// Mitsubishi GX Works2 project: 20国轩1次注液出1031   PLC: Q06UDEH

TYPE ConveyorIO : STRUCT
  xUnloadCCW : BOOL;  (* 下料为反转 *)
  xUnloadAlarm : BOOL;  (* 下料报警 *)
  xUnload : BOOL;  (* 下料请求 *)
  xPutInto : BOOL;  (* 线体直接投入物料 *)
  xNotArriveAlarm : BOOL;  (* 未到达报警 *)
  xNextRun : BOOL;  (* 下段线体运行 *)
  xMotorCW : BOOL;  (* 电机正转 *)
  xMotorCCW : BOOL;  (* 电机反转 *)
  xManual : BOOL;  (* 手动 *)
  xloadCCW : BOOL;  (* 上料为反转 *)
  xLimitAlarrm : BOOL;  (* 限位报警 *)
  xLoad : BOOL;  (* 上料请求 *)
  xForward : BOOL;  (* 正转手动 *)
  xEmpty : BOOL;  (* 线体状态为空 *)
  xCWPresent : BOOL;  (* 正转检测有无传感器 *)
  xCCWPresent : BOOL;  (* 反转检测有无传感器 *)
  xBusy : BOOL;  (* 工作中 *)
  xBackward : BOOL;  (* 反转手动 *)
  xAuto : BOOL;  (* 自动 *)
  xPosLimit : BOOL;  (* 正限位 *)
  xNegLimit : BOOL;  (* 负限位 *)
  xOverWidthAlarm : BOOL;  (* 超宽报警 *)
  xError : BOOL;  (* 报警 *)
  iProductCategoryIn : INT;  (* 产品类型输入 *)
  iProductCategory : INT;  (* 产品类型记录 *)
  iProductCategoryOut : INT;  (* 产品类型输出 *)
  diDeviceID : DINT;  (* 设备编号 *)
  tUnloadAlarmDelay : TIME;  (* 下料报警时间设置 *)
  tLoadDelay : TIME;  (* 上料延时设置 *)
  xSizeDeficientDetect : BOOL;  (* 尺寸缺陷检测 *)
  xZoneClear : BOOL;  (* 初始化线体清除 *)
  tZoneClearTime : TIME;  (* 初始化线体清除时间 *)
  iTaskIDIn : INT;  (* 产品类型输入 *)
  iTaskID : INT;  (* 产品类型记录 *)
  iTaskIDOut : INT;  (* 产品类型输出 *)
  diDesConveyorIn : DINT;  (* 产品类型输入 *)
  diDesConveyor : DINT;  (* 产品类型记录 *)
  diDesConveyorOut : DINT;  (* 产品类型输出 *)
END_STRUCT END_TYPE

TYPE QueueElement : STRUCT
  xCondition : BOOL;
  iPriority : INT;
END_STRUCT END_TYPE

TYPE ShuttleCarIO : STRUCT
  xReady : BOOL;  (* 准备就绪 *)
  xForward : BOOL;  (* 正转 *)
  xBackward : BOOL;  (* 反转 *)
  iCurrentPos : INT;  (* 当前位置 *)
  iDestinationPos : INT;  (* 目标位置 *)
  xCW : BOOL;  (* 正转输出 *)
  xCCW : BOOL;  (* 反转输出 *)
  xBrake : BOOL;  (* 刹车 *)
  xHomeSwitch : BOOL;  (* 零位接近开关 *)
  xPosLimit : BOOL;  (* 正限位 *)
  xNegLimit : BOOL;  (* 负限位 *)
  xMDIExe : BOOL;  (* MDI开始 *)
  xMDIDone : BOOL;  (* MDI 完成 *)
  xPassLimit : BOOL;  (* 限位屏蔽 *)
  xPosLimitCatch : BOOL;  (* 正限位捕捉 *)
  xNegLimitCatch : BOOL;  (* 负限位捕捉 *)
  xHomeExe : BOOL;  (* 开始寻零 *)
  xHomeDone : BOOL;  (* 寻零完成 *)
  xHomeBusy : BOOL;  (* 寻零中 *)
  xHomeFailed : BOOL;  (* 寻零失败 *)
  xBusy : BOOL;  (* 工作中 *)
  tArriveDelay : TIME;  (* 到位延时 *)
  xCylinder : BOOL;  (* 气缸控制 *)
  tBrakeDelay : TIME;  (* 抱闸延时 *)
  xPauseRamp : BOOL;  (* 暂停减速斜坡标志位 *)
  xPresentDetect1 : BOOL;  (* 物料有无检测1 *)
  xPresentDetect2 : BOOL;  (* 物料有无检测2 *)
  xOvertimeAlarm : BOOL;  (* 超时报警 *)
  tSetOverTime : TIME;  (* 设置超时时间 *)
  xLooseDetect : BOOL;  (* 松绳检测 *)
  xLooseAlarm : BOOL;  (* 松绳报警 *)
  xArrive : BOOL;  (* 到位信号 *)
  diDeviceID : DINT;  (* 设备编号 *)
  xMoveStep : BOOL;  (* 寸动 *)
  xAdrSwitch : ARRAY [1..8] OF BOOL;  (* 位置开关 *)
END_STRUCT END_TYPE

TYPE SwitchIO : STRUCT
  xLiftCylinderRetractDetect : BOOL;
  xLiftCylinderExtendDetect : BOOL;
  xLiftCylinderRetract : BOOL;
  xLiftCylinderExtend : BOOL;
  xEntryBarCylinderRetract : BOOL;
  xLiftCylinderExtendInit : BOOL;
  xEntryEnable : BOOL;
  xExitEnable : BOOL;
  xExitBarCylinderRetract : BOOL;
  xSwithEnable : BOOL;
  xLiftCylinderRetractButton : BOOL;
  xLiftCylinderExtendButton : BOOL;
  xEntryBarCylinderRetractButton : BOOL;
  xExitBarCylinderRetractButton : BOOL;
  xPutInto : BOOL;  (* 单体复位 *)
  tSetOvertime : TIME;  (* 设定超时报警时间 *)
  xOvertimeAlarm : BOOL;  (* 超时报警 *)
END_STRUCT END_TYPE

TYPE UConveyorIO : STRUCT
  xLiftCylinderRetractDetect1 : BOOL;
  xLiftCylinderRetractDetect2 : BOOL;
  xLiftCylinderExtendDetect1 : BOOL;
  xLiftCylinderExtendDetect2 : BOOL;
  xLiftCylinderRetract1 : BOOL;
  xLiftCylinderRetract2 : BOOL;
  xLiftCylinderExtend1 : BOOL;
  xLiftCylinderExtend2 : BOOL;
  xExitBarCylinderRetract1 : BOOL;
  xExitBarCylinderRetract2 : BOOL;
  xLiftCylinderExtendInit1 : BOOL;
  xLiftCylinderExtendInit2 : BOOL;
  xEntryEnable1 : BOOL;
  xEntryEnable2 : BOOL;
  xEntryEnable3 : BOOL;
  xExitEnable1 : BOOL;
  xExitEnable2 : BOOL;
  xExitEnable3 : BOOL;
  xPassEnable : BOOL;  (* 直接放行去下段 *)
  xLiftCylinderRetractButton1 : BOOL;
  xLiftCylinderRetractButton2 : BOOL;
  xLiftCylinderExtendButton1 : BOOL;
  xLiftCylinderExtendButton2 : BOOL;
  xExitBarCylinderRetractButton1 : BOOL;
  xExitBarCylinderRetractButton2 : BOOL;
  xPutInto : BOOL;  (* 单体复位 *)
  tSetOvertime : TIME;  (* 设定超时报警时间 *)
  xOvertimeAlarm : BOOL;  (* 超时报警 *)
  iTask : INT;  (* 3个任务 *)
  xBatteryDetect1 : BOOL;  (* 电池检测1 *)
  xBatteryDetect2 : BOOL;  (* 电池检测2 *)
  xBatteryError : BOOL;  (* 空框里有电池错误 *)
END_STRUCT END_TYPE

TYPE FanucRobotIO : STRUCT
  i_xCMDENBL : BOOL;
  i_xSYSRDY : BOOL;
  i_xPROG_RUN : BOOL;  (* 程序运行中 *)
  i_xPAUSED : BOOL;
  i_xHELD : BOOL;
  i_xFAULT : BOOL;
  i_xATPERCH : BOOL;
  i_xTPENBL : BOOL;
  i_xBATALM : BOOL;
  i_xBUSY : BOOL;  (* 工作中信号 *)
  i_arrxSNO : ARRAY [0..7] OF BOOL;  (* 传回的数据 *)
  i_xSNACK : BOOL;  (* 数据传回校验标志位 *)
  o_xIMSTP : BOOL;
  o_xHOLD : BOOL;
  o_xSFSPD : BOOL;
  o_xCSTOPI : BOOL;
  o_xRESET : BOOL;
  o_xSTART : BOOL;
  o_xENBL : BOOL;
  o_iPNS : INT;  (* 发给他的动作编号 *)
  o_xPNSTROBE : BOOL;  (* 传递动作编号标志位 *)
  o_xPROD_START : BOOL;  (* 启动信号，下降沿开动 *)
  o_xREMOTE : BOOL;  (* 远程模式开启 *)
  i_xCommandStart : BOOL;  (* 启动 *)
  i_iMotionNumber : INT;  (* 我程序给的动作编号 *)
  o_xPNSFailed : BOOL;  (* 程序号传输错误 *)
  o_uiOffset_X : INT;  (* X轴偏移量 *)
  o_uiOffset_Y : INT;  (* Y轴偏移量 *)
  io_xMutexLock : BOOL;  (* 互斥锁 *)
END_STRUCT END_TYPE

TYPE CommunicationIO : STRUCT
  i_iResponsPCPLC : INT;  (* 上位机写入-请求确认 *)
  i_iReadWriteFlagPCPLC : INT;  (* 上位机写入-读写标志位 *)
  i_iTaskProcessFlagPCPLC : INT;  (* 上位机写入-任务出料标志位 *)
  i_iCommandPCPLC : INT;  (* 上位机写入-命令字 *)
  i_iTaskIDPCPLC : INT;  (* 上位机写入-任务号 *)
  i_diDestinationDevicePCPLC : DINT;  (* 上位机写入-目标设备号 *)
  i_iProductIDPCPLC : INT;  (* 上位机写入-框码后4位 *)
  o_iRequestPLCPC : INT;  (* 上位机读取-请求状态 *)
  o_iReadWriteFlagPLCPC : INT;  (* 上位机读取-读写标志位 *)
  o_iDeviceStatusPLCPC : INT;  (* 上位机读取-设备状态 *)
  o_iTaskIDPLCPC : INT;  (* 上位机读取-任务号 *)
  o_iProductIDPLCPC : INT;  (* 上位机读取-框码后4位 *)
END_STRUCT END_TYPE

TYPE PackCommunicationIO : STRUCT
  i_iResponsPCPLC : INT;  (* 上位机写入-请求确认 *)
  i_iPackDoneAknPCPLC : INT;  (* 上位机写入-放行 *)
  i_iSinglePackResponsePCPLC : INT;  (* 上位机写入-单次装载应答 *)
  i_iSinglePackDoneAknPCPLC : INT;  (* 上位机写入-单次装载处理完成 *)
  o_iRequestPLCPC : INT;  (* 上位机读取-装载请求 *)
  o_iPackDonePLCPC : INT;  (* 上位机读取-装载完成 *)
  o_iSinglePackRequestPLCPC : INT;  (* 上位机读取-单次装载请求 *)
  o_iSinglePackDonePLCPC : INT;  (* 上位机读取-单次装载完成 *)
  o_iXCoordinatePLCPC : INT;  (* 上位机读取-行坐标 *)
  o_iYCoordinatePLCPC : INT;  (* 上位机读取-列坐标 *)
  o_arrwCode : ARRAY [0..7] OF BOOL;  (* 上位机读取-电芯码 *)
END_STRUCT END_TYPE

TYPE BatteryCode : STRUCT
  arrwCode : ARRAY [0..8] OF WORD;
END_STRUCT END_TYPE

// global labels: Global
VAR_GLOBAL
  g_xAuto AT M11 : BOOL;
  g_xManual : BOOL;
  g_xEStop AT X0 : BOOL;
  g_xReset AT X4 : BOOL;
  g_xStackLampRed AT Y200 : BOOL;
  g_xStackLampAmber AT Y201 : BOOL;
  g_xStackLampGreen AT Y202 : BOOL;
  g_xBuzzer AT Y203 : BOOL;
  g_xStop AT X3 : BOOL;
  g_xAutoStart AT X2 : BOOL;
  g_xRemoteAutoStart AT M0 : BOOL;
  g_xRemoteAuto AT M10 : BOOL;
  g_iState AT D40 : INT;
  g_iLocalAutoStep : BOOL;
  g_xAlarm : BOOL;
  g_xPause AT M3 : BOOL;  (* 暂停 *)
  g_diDeviceIDSelect AT D0 : DINT;
  g_xResetSingle AT M4 : BOOL;  (* 单线体复位 *)
  g_xInsertTask AT M5 : BOOL;  (* 插入任务 *)
  g_iInsertTaskID AT D2 : INT;  (* 插入任务号 *)
  g_iConveyorStatus AT D4 : INT;
  g_iInsertCategory AT D6 : INT;
  g_diInsertDesConveyor AT D8 : DINT;
  g_xTcpFailed : BOOL;
  g_xPickOver : ARRAY [1..4] OF BOOL;  (* 注液机给我们的信号，待定 *)
  g_xRobot1BatteryDetect : ARRAY [1..8] OF BOOL;
  g_xRobot2BatteryDetect : ARRAY [1..8] OF BOOL;
  g_xRobot3BatteryDetect : ARRAY [1..8] OF BOOL;
  g_xRobot4BatteryDetect : ARRAY [1..8] OF BOOL;
  g_xAutoLamp AT Y204 : BOOL;
  g_xAutoSwitch AT X1 : BOOL;
  g_xMute : BOOL;
  g_iLoadTask AT D50 : ARRAY [0..13] OF INT;
  g_xResetTask1 AT M9 : BOOL;  (* 复位排队任务的 *)
END_VAR

// global labels: Pro
VAR_GLOBAL
  g_xRobot1Pos1Done AT X0A0 : BOOL;  (* 机器人1工位1码垛完成 *)
  g_xRobot1Pos1Ready AT Y230 : BOOL;  (* 机器人1工位1空托盘到位 *)
  g_xRobot1Pos2Done AT X0A1 : BOOL;  (* 机器人1工位2码垛完成 *)
  g_xRobot1Pos2Ready AT Y231 : BOOL;  (* 机器人1工位2空托盘到位 *)
  g_xRobot2Pos1Done AT X0A2 : BOOL;  (* 机器人2工位1码垛完成 *)
  g_xRobot2Pos1Ready AT Y237 : BOOL;  (* 机器人2工位1空托盘到位 *)
  g_xRobot2Pos2Done AT X0A3 : BOOL;  (* 机器人2工位2码垛完成 *)
  g_xRobot2Pos2Ready AT Y239 : BOOL;  (* 机器人2工位2空托盘到位 *)
  g_xRobot3Pos1Done AT X0A4 : BOOL;  (* 机器人3工位1码垛完成 *)
  g_xRobot3Pos1Ready AT Y232 : BOOL;  (* 机器人3工位1空托盘到位 *)
  g_xRobot3Pos2Done AT X0A5 : BOOL;  (* 机器人3工位2码垛完成 *)
  g_xRobot3Pos2Ready AT Y233 : BOOL;  (* 机器人3工位2空托盘到位 *)
  g_xRobot4Pos1Done AT X0A6 : BOOL;  (* 机器人4工位1码垛完成 *)
  g_xRobot4Pos1Ready : BOOL;  (* 机器人4工位1空托盘到位 *)
  g_xRobot4Pos2Done AT X0A7 : BOOL;  (* 机器人4工位2码垛完成 *)
  g_xRobot4Pos2Ready : BOOL;  (* 机器人4工位2空托盘到位 *)
END_VAR

// task Task_01 (event TRUE, interval 0, priority 31): POU, TCP, START

FUNCTION_BLOCK Conveyor
VAR
  m_xPresentDelay : BOOL;  (* 有无判断延时 *)
  m_xLoadDelayOut : BOOL;  (* 上料延时输出 *)
  m_xInitial : BOOL;  (* 初始化 *)
  m_tUnloadTimer : TIME;  (* 下料计时器 *)
  m_tPresentDelayCurrentTime : TIME;
  m_tonUnloadAlam : TON;  (* 下料报警定时器 *)
  m_tonPresentDelay : TON;  (* 物料有无判断延时，防止误动作 *)
  m_tonNotArriveAlarm : TON;  (* 未到达报警计时 *)
  m_tonLoadDelay : TON;  (* 上料延时 *)
  m_tNotArriveCurrentTime : TIME;  (* 未到达报警计时当前时间 *)
  m_tLoadTimer : TIME;  (* 上料计时器 *)
  iStep : INT;  (* 上料步骤 *)
  m_wStateWord : INT;
END_VAR
VAR_IN_OUT
  ConveyorMotor : ConveyorIO;  (* 输送线输入输出 *)
END_VAR
VAR
  m_tonZoneClear : TON;  (* 初始化清除 *)
  m_tZoneClearCurrentTime : TIME;  (* 初始化清除当前时间 *)
  m_xAutoClear : BOOL;  (* 初始化清除标志位 *)
  m_xZoneClearDone : BOOL;  (* 初始化清除完成 *)
END_VAR
(*////////////////////////////////////////////////////////////////////////////////////////////////////////////
//传输线控制FB块，可控制单方向线体，双向旋转线体，支持双向上下料            
//线体初始化后为空的情况下输入xLoad信号即可进行上料动作，使用xLoadCCW信号可反方向上料
//增加了产品信息和产品种类的储存，当传输线为空和上料进行标志位为零的情况下清除产品信息和产品种类
//使用方式是在置位xLoad信号后，把产品信息和产品种类传入，等下料后自动清零
//线体不为空的情况下使用xUnload信号可进行下料动作，物料有无传感器的下降沿后出发计时器，延时断开传输线旋转
//单方向传输线体把xLoadCCW、xUnloadCCW设置为零，双向线体上料方向和下料反向的,方向固定的 把xUnloadCCW设置为1
//双方向线体双向都能上下料的要根据上料的方向来设置xLoadCCW,xUnloadCCW
//增加工作中信号xBusy当电机正转 显示为工作中
//增加上下料超时报警，xLoadAlarm，xUnloadAlarm，设定时间在LOAD_UNLOAD_TIME常量上，现在设置的为30秒
//增加xPutInto信号，用于直接投入的物料，检测开关感应到后，直接进入下料流程，上升沿有效
//离开延时改为变量 iLeaveDelay 默认为0 离开检测开关离输送线尾端比较远的线体需要根据情况设定100ms为单位
//增加初始化标志位，增加进入延时时间，初始化为进入延时时间为0 ，离开延时时间为2S，通过外围接口可以更改
//修改信息  修改后请增加版本
//12-17进行了优化，增加了未到达报警，当物料未传送到下一设备，就报未到达报警，使用xNextRun标志位制作，没有正常到达
//第0步，不能跳转到第一步把标志位复位，即出现中断情况，2秒后报警
//修改信息  修改后请增加版本
//上料延时增加为50ms防止干扰信号
//nextrun信号在 第三步也要复位
//增加限位报警
//增加超宽报警
//增加产品型号输出在下料的时候把产品型号输送给下一段线体
//增加线体单独复位
//增加任务插入功能配合全局变量
//增加暂停功能
//增加线体状态字显示  0 空闲 1：有料  2 工作中  3  超限报警 4 超宽报警  5 未到达报警  6 下料超时报警
//空料判断放在自动前，进行有无报警判断，然后跳转
//修改超限报警，与尺寸检测报警
////YAO      V1.0
//把所有的IF语句去掉，  IF语句占用指针存储区，容易造成存储区不足的现象
////YAO      V1.1
//初始化清除线体标志位xZoneClear
//ZPA zero pressure accumulation  Term that describes the Conveyor controls and mechanical scheme that will 
//cause loads to queue on a conveyor in discrete zones such that loads do not touch each other(wrapped boxed tray tote carton)
//除了产品信息外，还增加了目标地址，任务类型的数据传递。
//YAO      V1.0
///////////////////////////////////////////////////////////////////////////////////////////////////////////
(*********************************************************)
(*//初始化，
//上料延时位0S，下料报警延时为30S
//下料延时设一个比较大的时间，主要依靠xunload标志位来停止输送线，特殊情况可以用延时来停止物流线下料
//设置时间大的时候计时器会失效*)
IF NOT m_xInitial THEN
	ConveyorMotor.tLoadDelay:=T#100ms;
	ConveyorMotor.tUnloadAlarmDelay:=T#30s;
	ConveyorMotor.xPosLimit:=1;
	ConveyorMotor.xNegLimit:=1;
	ConveyorMotor.xSizeDeficientDetect:=0;
	ConveyorMotor.xZoneClear:=0;
	ConveyorMotor.tZoneClearTime:=T#10s;
	m_xInitial:=1;
END_IF;
(*//自动
//复位信号把步号置0，但xLoad与xUnload没有复位，调用程序需要注意复位后把这两个信号置零，以免发生误动作
//物料有无判断增加延时，防止开自动瞬间误动作发生*)
m_tonPresentDelay(IN:= ConveyorMotor.xCWPresent OR ConveyorMotor.xCCWPresent,
 PT:=T#100ms,
 Q:= m_xPresentDelay,
 ET:= m_tPresentDelayCurrentTime);
CASE iStep OF
0:(*//初始化*)
	ConveyorMotor.xMotorCW:=0;
	ConveyorMotor.xMotorCCW:=0;
	ConveyorMotor.xNextRun:=0;
	ConveyorMotor.iProductCategoryOut:=0;
	ConveyorMotor.iTaskIDOut:=0;
	ConveyorMotor.diDesConveyorOut:=0;
	out(NOT m_xPresentDelay,ConveyorMotor.xEmpty);(*	//判断物料有无传感器*)	
	mov(m_xPresentDelay AND g_xAuto AND NOT ConveyorMotor.xError,3,iStep);(*//自动情况下进行跳转*)(*无超限报警*)
	mov(NOT m_xPresentDelay AND g_xAuto AND NOT ConveyorMotor.xError,1,iStep);
1: (*//上料*)
	rst(ConveyorMotor.xLoad ,ConveyorMotor.iProductCategory);(*//上料开始清除产品信息*)
	rst(ConveyorMotor.xLoad ,ConveyorMotor.iTaskID);
	rst(ConveyorMotor.xLoad ,ConveyorMotor.diDesConveyor);
	mov(ConveyorMotor.xLoad,2,iStep);
2: (*//上料完成*)
	ConveyorMotor.iProductCategory:=ConveyorMotor.iProductCategoryIn;(* //产品信息传入*)
	ConveyorMotor.iTaskID:=ConveyorMotor.iTaskIDIn;
	ConveyorMotor.diDesConveyor:=ConveyorMotor.diDesConveyorIn;
	set(ConveyorMotor.xloadCCW,ConveyorMotor.xMotorCCW);
	rst(ConveyorMotor.xloadCCW,ConveyorMotor.xMotorCW);
	set(NOT ConveyorMotor.xloadCCW,ConveyorMotor.xMotorCW);
	rst(NOT ConveyorMotor.xloadCCW,ConveyorMotor.xMotorCCW);	
	m_tonLoadDelay(IN:= (ConveyorMotor.xCWPresent AND NOT ConveyorMotor.xloadCCW) 
  		OR (ConveyorMotor.xCCWPresent AND ConveyorMotor.xloadCCW) ,
  PT:= ConveyorMotor.tLoadDelay ,
  Q:= m_xLoadDelayOut ,
  ET:= m_tLoadTimer );
	mov(m_xLoadDelayOut,3, iStep);
3:(*//下料请求*)	
	ConveyorMotor.xMotorCW:=0;
	ConveyorMotor.xMotorCCW:=0;
	ConveyorMotor.xEmpty:=0;
	mov(ConveyorMotor.xUnload AND NOT ConveyorMotor.xOverWidthAlarm,4,iStep);
4:(*	//下料完成*)
	set(ConveyorMotor.xUnloadCCW,ConveyorMotor.xMotorCCW);
	rst(ConveyorMotor.xUnloadCCW,ConveyorMotor.xMotorCW);
	set(NOT ConveyorMotor.xUnloadCCW,ConveyorMotor.xMotorCW);
	rst(NOT ConveyorMotor.xUnloadCCW,ConveyorMotor.xMotorCCW);	
	ConveyorMotor.xNextRun:=1; (*下一段线体旋转*)
	ConveyorMotor.iProductCategoryOut:=ConveyorMotor.iProductCategory;(*产品型号输出给下一段线体*)
	ConveyorMotor.iTaskIDOut:=ConveyorMotor.iTaskID;
	ConveyorMotor.diDesConveyorOut:=ConveyorMotor.diDesConveyor;
	mov( NOT ConveyorMotor.xUnload , 0, istep );
END_CASE;
(*In-feed zone clear and ready to accept a load from upstream Conveyor*)
set(ldp(TRUE,g_xAuto) ,m_xAutoClear);
rst(ldf(TRUE,g_xAuto) ,m_xAutoClear);
m_tonZoneClear(IN:= m_xAutoClear AND ConveyorMotor.xZoneClear ,PT:= ConveyorMotor.tZoneClearTime ,Q:=m_xZoneClearDone ,ET:= m_tZoneClearCurrentTime );
set(m_xAutoClear AND ConveyorMotor.xZoneClear,ConveyorMotor.xMotorCW);
mov( m_xAutoClear AND ConveyorMotor.xZoneClear, 0 ,iStep );
rst(  ldf(TRUE, m_xAutoClear ) ,ConveyorMotor.xMotorCW);
rst( m_xZoneClearDone OR m_xPresentDelay  , m_xAutoClear );
(*投入上料，搬出下料，也可用来初始化*)
movp( ConveyorMotor.xPutInto, 0 , iStep );
(*//当前任务显示*)
movp( ConveyorMotor.diDeviceID=g_diDeviceIDSelect , ConveyorMotor.iProductCategory , g_iInsertCategory );
movp( ConveyorMotor.diDeviceID=g_diDeviceIDSelect , ConveyorMotor.iTaskID , g_iInsertTaskID );
dmovp( ConveyorMotor.diDeviceID=g_diDeviceIDSelect , ConveyorMotor.diDesConveyor , g_diInsertDesConveyor );
(*//插入任务*)
mov(g_xInsertTask AND ConveyorMotor.diDeviceID=g_diDeviceIDSelect ,g_iInsertCategory , ConveyorMotor.iProductCategory );
mov(g_xInsertTask AND ConveyorMotor.diDeviceID=g_diDeviceIDSelect , g_iInsertTaskID , ConveyorMotor.iTaskID );
dmov(g_xInsertTask AND ConveyorMotor.diDeviceID=g_diDeviceIDSelect , g_diInsertDesConveyor , ConveyorMotor.diDesConveyor );
(*//单线体复位，当设备号与本线体一致的时候执行复位*)
mov(g_xResetSingle AND ConveyorMotor.diDeviceID=g_diDeviceIDSelect , 0 , iStep );
rst(g_xResetSingle AND ConveyorMotor.diDeviceID=g_diDeviceIDSelect ,ConveyorMotor.xNextRun );
rst(g_xResetSingle AND ConveyorMotor.diDeviceID=g_diDeviceIDSelect  ,ConveyorMotor.xLimitAlarrm );
rst(g_xResetSingle AND ConveyorMotor.diDeviceID=g_diDeviceIDSelect  ,ConveyorMotor.xOverWidthAlarm );
(*//手动*)
(*//正转*)
set( g_xManual 
AND ConveyorMotor.xForward 
AND ConveyorMotor.xBackward=0 
AND ConveyorMotor.xMotorCCW=0 
AND g_xEStop  , 
ConveyorMotor.xMotorCW);
rst((g_xManual 
AND (NOT ConveyorMotor.xForward  
OR ConveyorMotor.xBackward 
OR ConveyorMotor.xMotorCCW )) 
OR  NOT g_xEStop,
ConveyorMotor.xMotorCW);
(*//反转*)		
set(g_xManual 
AND ConveyorMotor.xBackward 
AND ConveyorMotor.xForward=0 
AND ConveyorMotor.xMotorCW=0 
AND g_xEStop ,
ConveyorMotor.xMotorCCW);
rst((g_xManual AND 
(NOT ConveyorMotor.xBackward  
OR ConveyorMotor.xForward 
OR ConveyorMotor.xMotorCW ) ) 
OR NOT g_xEStop,
ConveyorMotor.xMotorCCW);
mov(g_xManual ,0,iStep);(*//手动后上下料程序步骤清零*)
(*暂停*)
rst(g_xPause,ConveyorMotor.xMotorCCW);
rst( g_xPause , ConveyorMotor.xMotorCW );
(*工作中信号输出*)
ConveyorMotor.xBusy:=ConveyorMotor.xMotorCCW OR ConveyorMotor.xMotorCW;
(*//未到达报警*)
m_tonNotArriveAlarm(IN:= iStep=0 AND ConveyorMotor.xNextRun  ,PT:= T#2s,Q:= ConveyorMotor.xNotArriveAlarm ,ET:= m_tNotArriveCurrentTime );
(*//下料超时报警*)
m_tonUnloadAlam(IN:= iStep=4,PT:=ConveyorMotor.tUnloadAlarmDelay,Q:= ConveyorMotor.xUnloadAlarm,ET:=m_tUnloadTimer );
(*//限位报警,进料检测开关失效*)
set(  ( ((ConveyorMotor.xloadCCW AND NOT ConveyorMotor.xNegLimit)            (*反转上料，碰到负限位*)
			OR  ( NOT ConveyorMotor.xloadCCW AND NOT ConveyorMotor.xPosLimit)) (*正转上料，碰到正限位*)
		AND iStep=2) (*上料过程*)
	OR
	( iStep=4 (*下料过程*)
		AND( (ConveyorMotor.xUnloadCCW AND NOT ConveyorMotor.xPosLimit)  
			OR (NOT ConveyorMotor.xUnloadCCW AND NOT ConveyorMotor.xNegLimit)))  ,  
	ConveyorMotor.xLimitAlarrm );
mov( ( ((ConveyorMotor.xloadCCW AND NOT ConveyorMotor.xNegLimit)            (*反转上料，碰到负限位*)
			OR  ( NOT ConveyorMotor.xloadCCW AND NOT ConveyorMotor.xPosLimit)) (*正转上料，碰到正限位*)
		AND iStep=2) (*上料过程*)
	OR
	( iStep=4 (*下料过程*)
		AND( (ConveyorMotor.xUnloadCCW AND NOT ConveyorMotor.xPosLimit)  
			OR (NOT ConveyorMotor.xUnloadCCW AND NOT ConveyorMotor.xNegLimit)))  ,
	0,
	iStep);
(*//超宽报警*)
set( (iStep=3 OR iStep=1) AND (NOT ConveyorMotor.xNegLimit OR NOT ConveyorMotor.xPosLimit) , ConveyorMotor.xOverWidthAlarm  );
(*//尺寸不足报警*)
(*//有料状态下检测两个开关都要有信号*)
set( iStep=3 AND ConveyorMotor.xSizeDeficientDetect AND (NOT ConveyorMotor.xCCWPresent OR NOT ConveyorMotor.xCWPresent) ,  ConveyorMotor.xOverWidthAlarm );
mov( iStep=3 AND ConveyorMotor.xSizeDeficientDetect AND (NOT ConveyorMotor.xCCWPresent OR NOT ConveyorMotor.xCWPresent),0,iStep);
(*//总报警*)
ConveyorMotor.xError:=ConveyorMotor.xLimitAlarrm
 OR ConveyorMotor.xNotArriveAlarm
 OR ConveyorMotor.xUnloadAlarm                                             
 OR ConveyorMotor.xOverWidthAlarm;

(*//状态输出*)(*状态显示，容易造成指针容量不足*)
mov( ConveyorMotor.xEmpty AND NOT ConveyorMotor.xBusy , 0 , m_wStateWord);
mov( ConveyorMotor.xEmpty=0 ,  		1 , m_wStateWord);
mov( ConveyorMotor.xBusy ,  			2 , m_wStateWord);
mov( ConveyorMotor.xLimitAlarrm ,  	3, 	m_wStateWord);
mov(ConveyorMotor.xOverWidthAlarm ,  4 , m_wStateWord);
mov( ConveyorMotor.xNotArriveAlarm ,  5 , m_wStateWord);
mov( ConveyorMotor.xUnloadAlarm,  	6 , m_wStateWord);
(*选择本线体后，将状态赋值给全局变量进行显示*)
mov( ConveyorMotor.diDeviceID=g_diDeviceIDSelect , m_wStateWord, g_iConveyorStatus );
END_FUNCTION_BLOCK

FUNCTION_BLOCK ConveyorOld
VAR
  m_xPresentDelay : BOOL;  (* 有无判断延时 *)
  m_xLoadDelayOut : BOOL;  (* 上料延时输出 *)
  m_xInitial : BOOL;  (* 初始化 *)
  m_tUnloadTimer : TIME;  (* 下料计时器 *)
  m_tPresentDelayCurrentTime : TIME;
  m_tonUnloadAlam : TON;  (* 下料报警定时器 *)
  m_tonPresentDelay : TON;  (* 物料有无判断延时，防止误动作 *)
  m_tonNotArriveAlarm : TON;  (* 未到达报警计时 *)
  m_tonLoadDelay : TON;  (* 上料延时 *)
  m_tNotArriveCurrentTime : TIME;  (* 未到达报警计时当前时间 *)
  m_tLoadTimer : TIME;  (* 上料计时器 *)
  iStep : INT;  (* 上料步骤 *)
  m_wStateWord : INT;
END_VAR
VAR_IN_OUT
  ConveyorMotor : ConveyorIO;  (* 输送线输入输出 *)
END_VAR
VAR
  m_tonZoneClear : TON;  (* 初始化清除 *)
  m_tZoneClearCurrentTime : TIME;  (* 初始化清除当前时间 *)
  m_xAutoClear : BOOL;  (* 初始化清除标志位 *)
  m_xZoneClearDone : BOOL;  (* 初始化清除完成 *)
END_VAR
(*////////////////////////////////////////////////////////////////////////////////////////////////////////////
//传输线控制FB块，可控制单方向线体，双向旋转线体，支持双向上下料            
//线体初始化后为空的情况下输入xLoad信号即可进行上料动作，使用xLoadCCW信号可反方向上料
//增加了产品信息和产品种类的储存，当传输线为空和上料进行标志位为零的情况下清除产品信息和产品种类
//使用方式是在置位xLoad信号后，把产品信息和产品种类传入，等下料后自动清零
//线体不为空的情况下使用xUnload信号可进行下料动作，物料有无传感器的下降沿后出发计时器，延时断开传输线旋转
//单方向传输线体把xLoadCCW、xUnloadCCW设置为零，双向线体上料方向和下料反向的,方向固定的 把xUnloadCCW设置为1
//双方向线体双向都能上下料的要根据上料的方向来设置xLoadCCW,xUnloadCCW
//增加工作中信号xBusy当电机正转 显示为工作中
//增加上下料超时报警，xLoadAlarm，xUnloadAlarm，设定时间在LOAD_UNLOAD_TIME常量上，现在设置的为30秒
//增加xPutInto信号，用于直接投入的物料，检测开关感应到后，直接进入下料流程，上升沿有效
//离开延时改为变量 iLeaveDelay 默认为0 离开检测开关离输送线尾端比较远的线体需要根据情况设定100ms为单位
//增加初始化标志位，增加进入延时时间，初始化为进入延时时间为0 ，离开延时时间为2S，通过外围接口可以更改
//修改信息  修改后请增加版本
//12-17进行了优化，增加了未到达报警，当物料未传送到下一设备，就报未到达报警，使用xNextRun标志位制作，没有正常到达
//第0步，不能跳转到第一步把标志位复位，即出现中断情况，2秒后报警
//修改信息  修改后请增加版本
上料延时增加为50ms防止干扰信号
nextrun信号在 第三步也要复位
增加限位报警
增加超宽报警
增加产品型号输出在下料的时候把产品型号输送给下一段线体
增加线体单独复位
增加任务插入功能配合全局变量
增加暂停功能
增加线体状态字显示  0 空闲 1：有料  2 工作中  3  超限报警 4 超宽报警  5 未到达报警  6 下料超时报警
空料判断放在自动前，进行有无报警判断，然后跳转
修改超限报警，与尺寸检测报警
初始化清除线体标志位xZoneClear
ZPA zero pressure accumulation  Term that describes the Conveyor controls and mechanical scheme that will 
cause loads to queue on a conveyor in discrete zones such that loads do not touch each other(wrapped boxed tray tote carton)
//YAO      V1.0
///////////////////////////////////////////////////////////////////////////////////////////////////////////
(*********************************************************)
(*//初始化，
//上料延时位0S，下料报警延时为30S
//下料延时设一个比较大的时间，主要依靠xunload标志位来停止输送线，特殊情况可以用延时来停止物流线下料
//设置时间大的时候计时器会失效*)
IF NOT m_xInitial THEN
	ConveyorMotor.tLoadDelay:=T#100ms;
	ConveyorMotor.tUnloadAlarmDelay:=T#30s;
	ConveyorMotor.xPosLimit:=1;
	ConveyorMotor.xNegLimit:=1;
	ConveyorMotor.xSizeDeficientDetect:=0;
	ConveyorMotor.xZoneClear:=0;
	ConveyorMotor.tZoneClearTime:=T#10s;
	m_xInitial:=1;
END_IF;
(*//自动
//复位信号把步号置0，但xLoad与xUnload没有复位，调用程序需要注意复位后把这两个信号置零，以免发生误动作
//物料有无判断增加延时，防止开自动瞬间误动作发生*)
m_tonPresentDelay(IN:= ConveyorMotor.xCWPresent OR ConveyorMotor.xCCWPresent,
                  PT:=T#100ms,
				  Q:= m_xPresentDelay,
				  ET:= m_tPresentDelayCurrentTime);

CASE iStep OF
	0:(*//初始化*)
	ConveyorMotor.xMotorCW:=0;
	ConveyorMotor.xMotorCCW:=0;
	ConveyorMotor.iProductCategoryOut:=0;
(*	//判断物料有无传感器*)	
		IF m_xPresentDelay THEN			
			ConveyorMotor.xEmpty:=0;
			IF g_xAuto AND NOT ConveyorMotor.xError THEN(*//自动情况下进行跳转*)(*无超限报警*)
				iStep:=3;
			END_IF;
		ELSE
			ConveyorMotor.xEmpty:=1;
			IF g_xAuto AND NOT ConveyorMotor.xError THEN(*//自动情况下进行跳转*)(*无超限报警*)
				iStep:=1;	
			END_IF;		
	END_IF;	
	1: (*//上料*)
	ConveyorMotor.xNextRun:=0;
	IF ConveyorMotor.xLoad    THEN (*//上料开始*)
		ConveyorMotor.iProductCategory:=0;	(*//上料开始清除产品信息*)
		iStep:=2;		
	END_IF;
	2: (*//上料完成*)
	IF ConveyorMotor.iProductCategoryIn<>0 THEN
		ConveyorMotor.iProductCategory:=ConveyorMotor.iProductCategoryIn;(* //产品信息传入*)
	END_IF;
	IF ConveyorMotor.xloadCCW THEN
		ConveyorMotor.xMotorCCW:=1; 
		ConveyorMotor.xMotorCW:=0;
	ELSE
	    ConveyorMotor.xMotorCW:=1;  
		ConveyorMotor.xMotorCCW:=0;
	END_IF;
		m_tonLoadDelay(IN:= (ConveyorMotor.xCWPresent AND NOT ConveyorMotor.xloadCCW) 
		                                        OR (ConveyorMotor.xCCWPresent AND ConveyorMotor.xloadCCW) ,
		                               PT:= ConveyorMotor.tLoadDelay ,
		                               Q:= m_xLoadDelayOut ,
		                               ET:= m_tLoadTimer );
	    IF m_xLoadDelayOut THEN 	 
		    iStep:=3;
		END_IF;
	3:(*//下料请求*)	
	ConveyorMotor.xMotorCW:=0;
	ConveyorMotor.xMotorCCW:=0;
	ConveyorMotor.xEmpty:=0;
	IF ConveyorMotor.xUnload AND NOT ConveyorMotor.xOverWidthAlarm  THEN (*无超宽报警可以下料*)
		iStep:=4;
	END_IF;
	4:(*	//下料完成*)
	IF ConveyorMotor.xUnloadCCW THEN   
		ConveyorMotor.xMotorCCW:=1;  
		ConveyorMotor.xMotorCW:=0;
		ELSE
	    ConveyorMotor.xMotorCW:=1;  
		ConveyorMotor.xMotorCCW:=0;
	END_IF;
	ConveyorMotor.xNextRun:=1; (*下一段线体旋转*)
	ConveyorMotor.iProductCategoryOut:=ConveyorMotor.iProductCategory;(*产品型号输出给下一段线体*)
	IF NOT ConveyorMotor.xUnload THEN 
		istep:=0;
	END_IF;
END_CASE;
(*In-feed zone clear and ready to accept a load from upstream Conveyor*)
IF ldp(TRUE,g_xAuto) THEN
	m_xAutoClear:=1;
END_IF;
IF ldf(TRUE,g_xAuto) THEN
	m_xAutoClear:=0;
END_IF;
m_tonZoneClear(IN:= m_xAutoClear AND ConveyorMotor.xZoneClear ,PT:= ConveyorMotor.tZoneClearTime ,Q:=m_xZoneClearDone ,ET:= m_tZoneClearCurrentTime );
IF  m_xAutoClear AND ConveyorMotor.xZoneClear THEN
		ConveyorMotor.xMotorCW:=1; 
		iStep:=0;
END_IF;
IF ldf(TRUE, m_xAutoClear )THEN
	ConveyorMotor.xMotorCW:=0; 
END_IF;
IF NOT m_xAutoClear OR m_xZoneClearDone OR m_xPresentDelay THEN
	 m_xAutoClear:=0;
END_IF;	 
(*投入上料，搬出下料，也可用来初始化*)
IF LDP(TRUE,ConveyorMotor.xPutInto) THEN
	iStep:=0;
END_IF;
(*//当前任务显示*)
IF LDP(TRUE,ConveyorMotor.iDeviceID=g_iDeviceIDSelect) THEN
	g_iInsertTask:=ConveyorMotor.iProductCategory;
END_IF;
	(*//插入任务*)
IF g_xInsertTask AND ConveyorMotor.iDeviceID=g_iDeviceIDSelect THEN
	ConveyorMotor.iProductCategory:=g_iInsertTask;
END_IF;
(*//单线体复位，当设备号与本线体一致的时候执行复位*)
IF (g_xResetSingle AND ConveyorMotor.iDeviceID=g_iDeviceIDSelect)THEN (* //非正常情况下切断xNextRun不会复位，通过这个标志位会出发报警*)(*增加单体复位*)
	iStep:=0;
	ConveyorMotor.xNextRun:=0; 
	ConveyorMotor.xLimitAlarrm:=0;
	ConveyorMotor.xOverWidthAlarm:=0;
END_IF;
(*//手动*)
IF g_xManual THEN
(*	iStep:=0; *)(*//手动后上下料程序步骤清零*)
	(*//正转*)
	IF ConveyorMotor.xForward 
		AND ConveyorMotor.xBackward=0 
		AND ConveyorMotor.xMotorCCW=0 
		AND g_xEStop THEN
		ConveyorMotor.xMotorCW:=1;
		ConveyorMotor.xMotorCCW:=0;
		ELSE
		ConveyorMotor.xMotorCW:=0;
	END_IF;
	(*//反转*)
	IF ConveyorMotor.xBackward 
		AND ConveyorMotor.xForward=0 
		AND ConveyorMotor.xMotorCW=0 
		AND g_xEStop THEN
		ConveyorMotor.xMotorCCW:=1;
		conveyormotor.xMotorCW:=0;
		ELSE
		ConveyorMotor.xMotorCCW:=0;
	END_IF;
END_IF;
(*暂停*)
IF g_xPause THEN
	ConveyorMotor.xMotorCCW:=0;
	ConveyorMotor.xMotorCW:=0;
END_IF;
(*工作中信号输出*)
ConveyorMotor.xBusy:=ConveyorMotor.xMotorCCW OR ConveyorMotor.xMotorCW;
(*//未到达报警*)
m_tonNotArriveAlarm(IN:= iStep=0 AND ConveyorMotor.xNextRun  ,PT:= T#2s,Q:= ConveyorMotor.xNotArriveAlarm ,ET:= m_tNotArriveCurrentTime );
(*//下料超时报警*)
m_tonUnloadAlam(IN:= iStep=4,PT:=ConveyorMotor.tUnloadAlarmDelay,Q:= ConveyorMotor.xUnloadAlarm,ET:=m_tUnloadTimer );
(*//限位报警,进料检测开关失效*)
IF ( ((ConveyorMotor.xloadCCW AND NOT ConveyorMotor.xNegLimit)            (*反转上料，碰到负限位*)
	OR  ( NOT ConveyorMotor.xloadCCW AND NOT ConveyorMotor.xPosLimit)) (*正转上料，碰到正限位*)
    AND iStep=2) (*上料过程*)
    OR
   ( iStep=4 (*下料过程*)
	AND( (ConveyorMotor.xUnloadCCW AND NOT ConveyorMotor.xPosLimit)  
	OR (NOT ConveyorMotor.xUnloadCCW AND NOT ConveyorMotor.xNegLimit)))    
    THEN
    ConveyorMotor.xLimitAlarrm:=1;
    iStep:=0;
END_IF;
(*//超宽报警*)
IF (iStep=3 OR iStep=1) AND (NOT ConveyorMotor.xNegLimit OR NOT ConveyorMotor.xPosLimit) THEN
	ConveyorMotor.xOverWidthAlarm:=1;
END_IF;
(*//尺寸不足报警*)
(*//有料状态下检测两个开关都要有信号*)
IF iStep=3 AND ConveyorMotor.xSizeDeficientDetect AND (NOT ConveyorMotor.xCCWPresent OR NOT ConveyorMotor.xCWPresent)  THEN
	   ConveyorMotor.xOverWidthAlarm:=1;
	    iStep:=0;               
END_IF;
(*//总报警*)
ConveyorMotor.xError:=ConveyorMotor.xLimitAlarrm
                                              OR ConveyorMotor.xNotArriveAlarm
                                              OR ConveyorMotor.xUnloadAlarm                                             
                                              OR ConveyorMotor.xOverWidthAlarm;

(*//状态输出*)(*状态显示，容易造成指针容量不足*)
IF ConveyorMotor.xEmpty AND NOT ConveyorMotor.xBusy THEN
	m_wStateWord:=0;
END_IF;
IF ConveyorMotor.xEmpty=0 THEN
		m_wStateWord:=1;
END_IF;
IF ConveyorMotor.xBusy THEN
		m_wStateWord:=2;
END_IF;
IF ConveyorMotor.xLimitAlarrm THEN
		m_wStateWord:=3;
END_IF;
IF ConveyorMotor.xOverWidthAlarm THEN
		m_wStateWord:=4;
END_IF;
IF ConveyorMotor.xNotArriveAlarm THEN	
		m_wStateWord:=5;
END_IF;
IF ConveyorMotor.xUnloadAlarm THEN
		m_wStateWord:=6;	
END_IF;
(*选择本线体后，将状态赋值给全局变量进行显示*)
IF ConveyorMotor.iDeviceID=g_iDeviceIDSelect THEN
	g_iConveyorStatus:=m_wStateWord;
END_IF;
END_FUNCTION_BLOCK

PROGRAM POU
VAR
  Conveyor20101 : Conveyor;
  Conveyor20102 : Conveyor;
  Conveyor20103 : Conveyor;
  Conveyor20104 : Conveyor;
  Conveyor20105 : Conveyor;
  Conveyor20106 : Conveyor;
  Conveyor20107 : Conveyor;
  Conveyor20108 : Conveyor;
  Conveyor20109 : Conveyor;
  Conveyor20110 : Conveyor;
  Conveyor20111 : Conveyor;
  Conveyor20112 : Conveyor;
  Conveyor20113 : Conveyor;
  Conveyor20114 : Conveyor;
  Conveyor20115 : Conveyor;
  Conveyor20116 : Conveyor;
  Conveyor20117 : Conveyor;
  Conveyor20118 : Conveyor;
  Conveyor20122 : Conveyor;
  Conveyor20123 : Conveyor;
  Conveyor20124 : Conveyor;
  Conveyor20125 : Conveyor;
  Conveyor20126 : Conveyor;
  Conveyor20127 : Conveyor;
  Conveyor20128 : Conveyor;
  Conveyor20129 : Conveyor;
  Conveyor20130 : Conveyor;
  Conveyor201021 : Conveyor;  (* 虚构的 *)
  Conveyor201031 : Conveyor;  (* 虚构的 *)
  Conveyor201041 : Conveyor;  (* 虚构的 *)
  Conveyor201051 : Conveyor;  (* 虚构的 *)
  Conveyor201061 : Conveyor;  (* 虚构的 *)
  Conveyor201071 : Conveyor;  (* 虚构的 *)
  Conveyor201081 : Conveyor;  (* 虚构的 *)
  Conveyor201091 : Conveyor;  (* 虚构的 *)
  ConveyorIO20101 : ConveyorIO;
  ConveyorIO20102 : ConveyorIO;
  ConveyorIO20103 : ConveyorIO;
  ConveyorIO20104 : ConveyorIO;
  ConveyorIO20105 : ConveyorIO;
  ConveyorIO20106 : ConveyorIO;
  ConveyorIO20107 : ConveyorIO;
  ConveyorIO20108 : ConveyorIO;
  ConveyorIO20109 : ConveyorIO;
  ConveyorIO20110 : ConveyorIO;
  ConveyorIO20111 : ConveyorIO;
  ConveyorIO20112 : ConveyorIO;
  ConveyorIO20113 : ConveyorIO;
  ConveyorIO20114 : ConveyorIO;
  ConveyorIO20115 : ConveyorIO;
  ConveyorIO20116 : ConveyorIO;
  ConveyorIO20117 : ConveyorIO;
  ConveyorIO20118 : ConveyorIO;
  ConveyorIO20122 : ConveyorIO;
  ConveyorIO20123 : ConveyorIO;
  ConveyorIO20124 : ConveyorIO;
  ConveyorIO20125 : ConveyorIO;
  ConveyorIO20126 : ConveyorIO;
  ConveyorIO20127 : ConveyorIO;
  ConveyorIO20128 : ConveyorIO;
  ConveyorIO20129 : ConveyorIO;
  ConveyorIO20130 : ConveyorIO;
  ConveyorIO201021 : ConveyorIO;  (* 虚构的 *)
  ConveyorIO201031 : ConveyorIO;  (* 虚构的 *)
  ConveyorIO201041 : ConveyorIO;  (* 虚构的 *)
  ConveyorIO201051 : ConveyorIO;  (* 虚构的 *)
  ConveyorIO201061 : ConveyorIO;  (* 虚构的 *)
  ConveyorIO201071 : ConveyorIO;  (* 虚构的 *)
  ConveyorIO201081 : ConveyorIO;  (* 虚构的 *)
  ConveyorIO201091 : ConveyorIO;  (* 虚构的 *)
  UConveyor20301 : UConveyor;
  UConveyor20303 : UConveyor;
  UConveyor20305 : UConveyor;
  UConveyor20307 : UConveyor;
  UConveyorIO20301 : UConveyorIO;
  UConveyorIO20303 : UConveyorIO;
  UConveyorIO20305 : UConveyorIO;
  UConveyorIO20307 : UConveyorIO;
  Switch20309 : Switch;
  Switch20312 : Switch;
  Switch20310 : Switch;
  Switch20311 : Switch;
  SwitchIO20309 : SwitchIO;
  SwitchIO20310 : SwitchIO;
  SwitchIO20311 : SwitchIO;
  SwitchIO20312 : SwitchIO;
  Conveyor201191 : Conveyor;  (* 虚构的 *)
  ConveyorIO201191 : ConveyorIO;  (* 虚构的 *)
  Lifter20201 : ShuttleCar;
  LifterIO20201 : ShuttleCarIO;
  Conveyor20101Task : PriorityQueue;  (* 上料排队任务 *)
  Conveyor20101Condition : ARRAY [1..13] OF QueueElement;  (* 上料排队任务 *)
  m_i20101Task : INT;  (* 上料排队任务 *)
  m_xLoadPermit : ARRAY [2..9] OF BOOL;
  Task20301 : PreemptivePriority;
  TaskCondition20301 : ARRAY [1..13] OF BOOL;
  Task20303 : PreemptivePriority;
  TaskCondition20303 : ARRAY [1..13] OF BOOL;
  Task20305 : PreemptivePriority;
  TaskCondition20305 : ARRAY [1..13] OF BOOL;
  Task20307 : PreemptivePriority;
  TaskCondition20307 : ARRAY [1..13] OF BOOL;
  m_xCatchCylinder : ARRAY [2..9] OF BOOL;
  ComConveyorIO30103 : CommunicationIO;
  ComConveyorIO20109 : CommunicationIO;
  ComConveyorIO20108 : CommunicationIO;
  ComConveyorIO20107 : CommunicationIO;
  ComConveyorIO20106 : CommunicationIO;
  ComConveyorIO20105 : CommunicationIO;
  ComConveyorIO20104 : CommunicationIO;
  ComConveyorIO20103 : CommunicationIO;
  ComConveyorIO20102 : CommunicationIO;
  ComConveyor30103 : ConveyorCommunication;
  ComConveyor20109 : ConveyorCommunication;
  ComConveyor20108 : ConveyorCommunication;
  ComConveyor20107 : ConveyorCommunication;
  ComConveyor20106 : ConveyorCommunication;
  ComConveyor20105 : ConveyorCommunication;
  ComConveyor20104 : ConveyorCommunication;
  ComConveyor20103 : ConveyorCommunication;
  ComConveyor20102 : ConveyorCommunication;
  Robot20901 : FanucRobot;
  Robot20902 : FanucRobot;
  Robot20903 : FanucRobot;
  Robot20904 : FanucRobot;
  RobotIO20901 : FanucRobotIO;
  RobotIO20902 : FanucRobotIO;
  RobotIO20903 : FanucRobotIO;
  RobotIO20904 : FanucRobotIO;
  PackCommunication20102 : PackCommunication;
  PackCommunication20103 : PackCommunication;
  PackCommunication20104 : PackCommunication;